(* Logix 5000 project; controller Seperator 1756-L85E rev 33.11; software revision 33.01; part 4 of 7 *)

ADD_ON_INSTRUCTION Random_Izer   (* revision 1.0 *)
VAR_IN_OUT
   Medium_Flash_ON : BOOL; {required}
   Energy : REAL; {required}
END_VAR
VAR_INPUT
   High_Limit_Reached : DINT;
   Actual_To_Same_Interval_Prior_Periods : REAL;
   Production_Lines_To_Like_Lines : REAL;
   Actual_to_Baseline : REAL;
   Production_Runs_To_Like_Runs : REAL;
   Eunits_PER_UOPunits : REAL;
   Edollar_PER_UOPunits : REAL;
   Eunits_PER_UOPdollar : REAL;
   Edollar_PER_UOPdollar : REAL;
   kG_CO2_e : REAL;
   Metric_Tonnes : REAL;
   Water_Demand : REAL;
   Air_Demand : REAL;
   Gas_Demand : REAL;
   Electric_Demand : REAL;
   Steam_Demand : REAL;
   Water_Usage : REAL;
   Air_Usage : REAL;
   Gas_Usage : REAL;
   Electric_Usage : REAL;
   Steam_Usage : REAL;
   work : REAL;
END_VAR
VAR
   APAC_ONS : DINT;
   Low_Limit_Reached : DINT;
   Enable_Low_Check : BOOL; {access None}
   Low_Limit : REAL := 20.0; {access None}
   High_Limit : REAL := 95.0; {access None}
   High_High_Limit : REAL := 100.0; {access None}
   Low_Low_Limit : REAL; {access None}
   Enable_Hi_Check : BOOL; {access None}
   ons1 : BOOL; {access None}
   ons2 : BOOL; {access None}
END_VAR

ROUTINE Logic   (* ladder *)
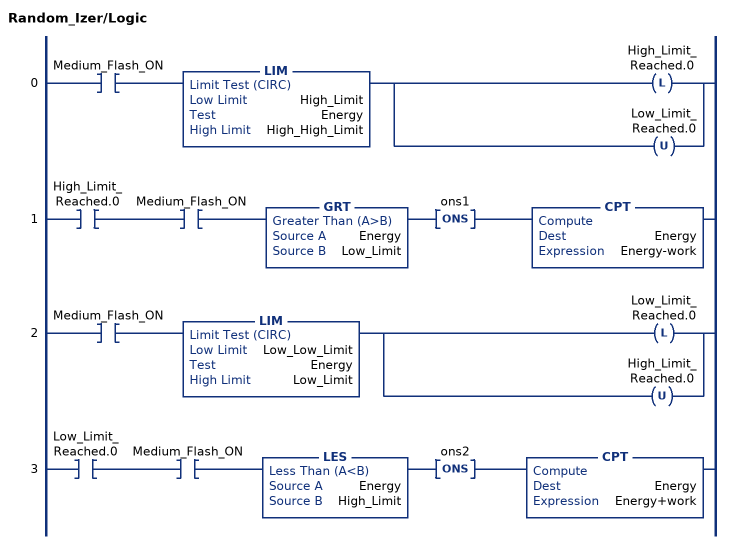
   0: XIC(Medium_Flash_ON)LIM(High_Limit,Energy,High_High_Limit)[OTL(High_Limit_Reached.0) ,OTU(Low_Limit_Reached.0) ];
   1: XIC(High_Limit_Reached.0)XIC(Medium_Flash_ON)GRT(Energy,Low_Limit)ONS(ons1)CPT(Energy,Energy-work);
   2: XIC(Medium_Flash_ON)LIM(Low_Low_Limit,Energy,Low_Limit)[OTL(Low_Limit_Reached.0) ,OTU(High_Limit_Reached.0) ];
   3: XIC(Low_Limit_Reached.0)XIC(Medium_Flash_ON)LES(Energy,High_Limit)ONS(ons2)CPT(Energy,Energy+work);
END_ROUTINE
END_ADD_ON_INSTRUCTION

ADD_ON_INSTRUCTION SineWave   (* revision 1.0, ExecutePrescan *)
VAR_INPUT
   Period : DINT; {visible}
   Max : REAL; {visible}
END_VAR
VAR_IN_OUT
   Out : INT; {required}
END_VAR
VAR
   PI : REAL;
   AlaFillerTimer : TIMER := (PRE := 20000, DN := 1);
   XNum : REAL;
   XDen : REAL;
   Ctrl : CONTROL := (LEN := 1);
   Ctrl2 : CONTROL;
END_VAR

ROUTINE Logic   (* ladder *)
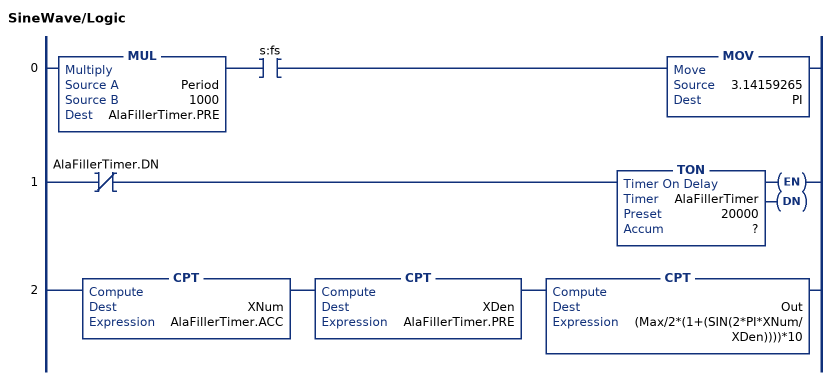
   0: MUL(Period,1000,AlaFillerTimer.PRE)XIC(s:fs)MOV(3.14159265,PI);
   1: XIO(AlaFillerTimer.DN)TON(AlaFillerTimer,?,?);
   2: CPT(XNum,AlaFillerTimer.ACC)CPT(XDen,AlaFillerTimer.PRE)CPT(Out,(Max/2*(1+(SIN(2*PI*XNum/XDen))))*10);
END_ROUTINE

ROUTINE Prescan   (* structured text *)
   Period:=20;
   Max:=50;
END_ROUTINE
END_ADD_ON_INSTRUCTION

ADD_ON_INSTRUCTION UADD   (* revision 1.1, vendor Dr. Frank Jordan / Rockwell Automation *)
// Addition of  two unsigned DINT
// (without overflow / minor faults)
// Revision note:
// This code is provided as application example without any warranty
VAR_INPUT
   V1 : DINT; {visible}
   V2 : DINT; {visible}
END_VAR
VAR_OUTPUT
   Out : DINT; {access Read Only, visible}
   Sts_C : BOOL; {access Read Only, visible}   // Carry result
   Sts_N : BOOL; {access Read Only, visible}   // Negative result
   Sts_V : BOOL; {access Read Only, visible}   // Overflow result
   Sts_Z : BOOL; {access Read Only, visible}   // Zero result
END_VAR
VAR
   V1_Hi : DINT; {access None}
   V1_Lo : DINT; {access None}
   V2_Hi : DINT; {access None}
   V2_Lo : DINT; {access None}
   SumLo : DINT; {access None}
   SumHi : DINT; {access None}
   tmp : DINT; {access None}
END_VAR

ROUTINE Logic   (* ladder *)
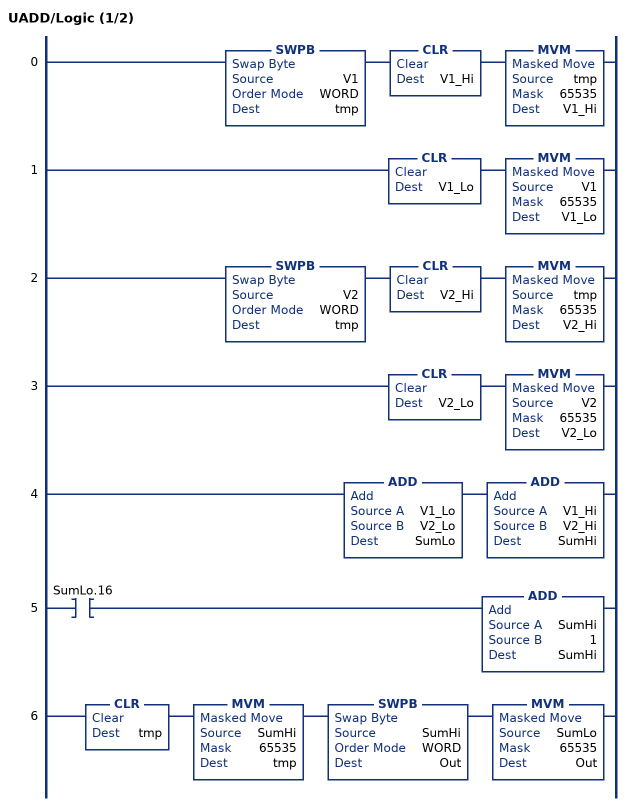
   0: SWPB(V1,WORD,tmp)CLR(V1_Hi)MVM(tmp,65535,V1_Hi);
   1: CLR(V1_Lo)MVM(V1,65535,V1_Lo);
   2: SWPB(V2,WORD,tmp)CLR(V2_Hi)MVM(tmp,65535,V2_Hi);
   3: CLR(V2_Lo)MVM(V2,65535,V2_Lo);
   4: ADD(V1_Lo,V2_Lo,SumLo)ADD(V1_Hi,V2_Hi,SumHi);
   5: XIC(SumLo.16)ADD(SumHi,1,SumHi);
   6: CLR(tmp)MVM(SumHi,65535,tmp)SWPB(SumHi,WORD,Out)MVM(SumLo,65535,Out);
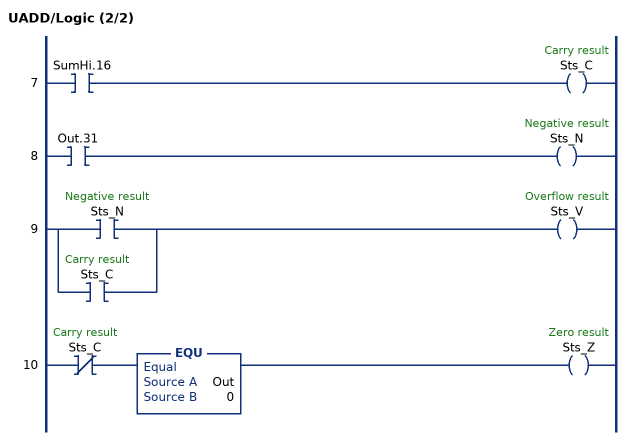
   7: XIC(SumHi.16)OTE(Sts_C);
   8: XIC(Out.31)OTE(Sts_N);
   9: [XIC(Sts_N) ,XIC(Sts_C) ]OTE(Sts_V);
   10: XIO(Sts_C)EQU(Out,0)OTE(Sts_Z);
END_ROUTINE
END_ADD_ON_INSTRUCTION

ADD_ON_INSTRUCTION UMUL   (* revision 1.2, vendor Dr. Frank Jordan / Rockwell Automation *)
// Multiplication of  two unsigned DINT
// (without overflow / minor faults)
// Revision note:
// This code is provided as application example without any warranty
VAR_INPUT
   V1 : DINT; {visible}
   V2 : DINT; {visible}
END_VAR
VAR_OUTPUT
   Sts_C : BOOL; {access Read Only, visible}   // Carry result
   Sts_N : BOOL; {access Read Only, visible}   // Negative result
   Sts_V : BOOL; {access Read Only, visible}   // Overflow result
   Sts_Z : BOOL; {access Read Only, visible}   // Zero result
   Out : DINT; {access Read Only, visible}
END_VAR
VAR
   tmp : DINT; {access None}
   WRK : INT[6]; {access None}
   WRKm : DINT[6]; {access None}
   Low : DINT; {access None}
   Mid : DINT; {access None}
   High : DINT; {access None}
END_VAR

ROUTINE Logic   (* ladder *)
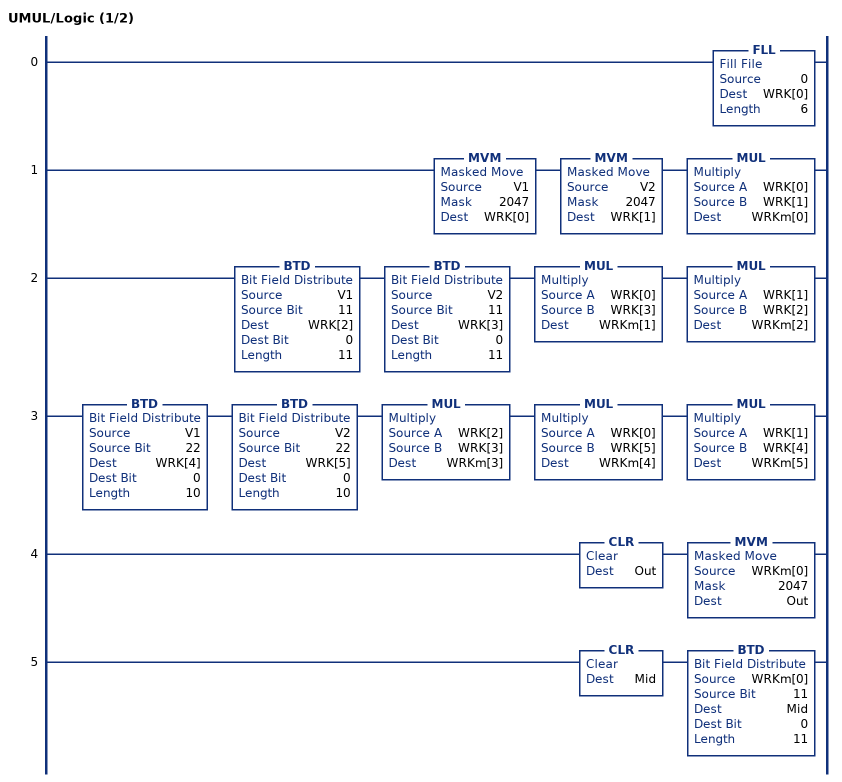
   0: FLL(0,WRK[0],6);
   1: MVM(V1,2047,WRK[0])MVM(V2,2047,WRK[1])MUL(WRK[0],WRK[1],WRKm[0]);
   2: BTD(V1,11,WRK[2],0,11)BTD(V2,11,WRK[3],0,11)MUL(WRK[0],WRK[3],WRKm[1])MUL(WRK[1],WRK[2],WRKm[2]);
   3: BTD(V1,22,WRK[4],0,10)BTD(V2,22,WRK[5],0,10)MUL(WRK[2],WRK[3],WRKm[3])MUL(WRK[0],WRK[5],WRKm[4])MUL(WRK[1],WRK[4],WRKm[5]);
   4: CLR(Out)MVM(WRKm[0],2047,Out);
   5: CLR(Mid)BTD(WRKm[0],11,Mid,0,11);
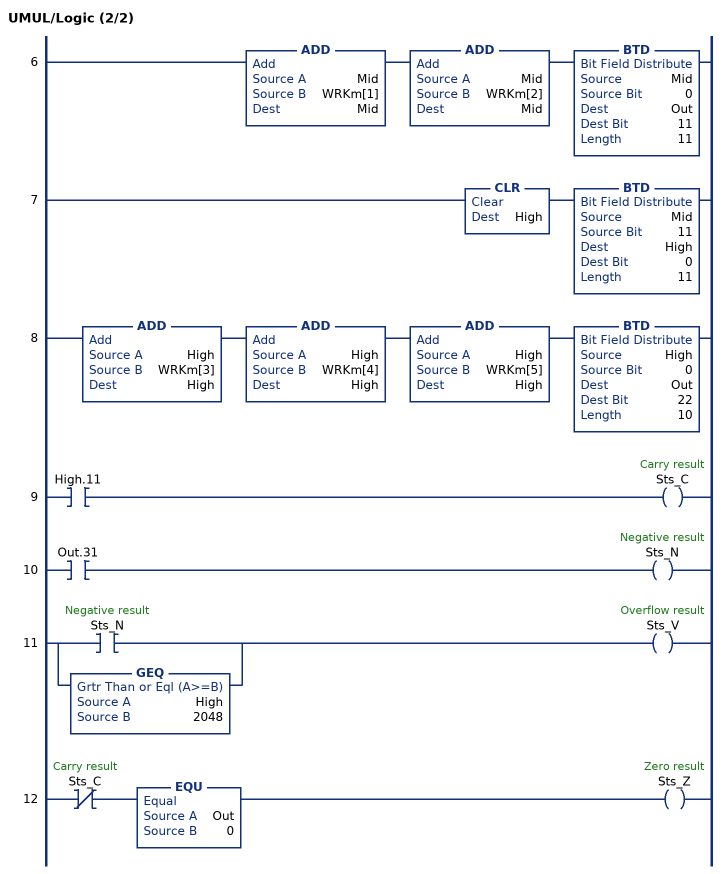
   6: ADD(Mid,WRKm[1],Mid)ADD(Mid,WRKm[2],Mid)BTD(Mid,0,Out,11,11);
   7: CLR(High)BTD(Mid,11,High,0,11);
   8: ADD(High,WRKm[3],High)ADD(High,WRKm[4],High)ADD(High,WRKm[5],High)BTD(High,0,Out,22,10);
   9: XIC(High.11)OTE(Sts_C);
   10: XIC(Out.31)OTE(Sts_N);
   11: [XIC(Sts_N) ,GEQ(High,2048) ]OTE(Sts_V);
   12: XIO(Sts_C)EQU(Out,0)OTE(Sts_Z);
END_ROUTINE
END_ADD_ON_INSTRUCTION

ADD_ON_INSTRUCTION ValveSim   (* revision 1.0, vendor Rockwell, ExecutePrescan *)
VAR_INPUT
   ValveOpenRequest : BOOL;
END_VAR
VAR_OUTPUT
   ValveOpened : BOOL; {access Read Only}
   ValveClosed : BOOL; {access Read Only}
END_VAR
VAR
   OpenCommand : BOOL;
   OpenedCommandDelay : TIMER := (PRE := 1000);
   ClosedCommandDelay : TIMER := (PRE := 1000);
END_VAR

ROUTINE Logic   (* ladder *)
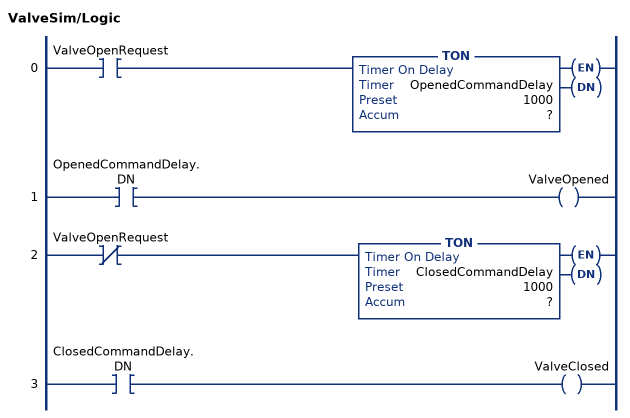
   0: XIC(ValveOpenRequest)TON(OpenedCommandDelay,?,?);
   1: XIC(OpenedCommandDelay.DN)OTE(ValveOpened);
   2: XIO(ValveOpenRequest)TON(ClosedCommandDelay,?,?);
   3: XIC(ClosedCommandDelay.DN)OTE(ValveClosed);
END_ROUTINE

ROUTINE Prescan   (* structured text *)
   OpenedCommandDelay.PRE:=3000;
   ClosedCommandDelay.PRE:=3000;
   
END_ROUTINE
END_ADD_ON_INSTRUCTION

VAR_GLOBAL   (* controller tags *)
   _DriveName_FP : BOOL;
   Aborted : SFC_STEP := (Status := 16#0020_0001, PauseTimer := 1);
   Aborted1 : SFC_STEP := (Status := 16#0020_0001, PauseTimer := 1);
   Aborting : SFC_STEP := (Status := 16#0020_0001, PauseTimer := 1);
   Aborting1 : SFC_STEP := (Status := 16#0020_0001, PauseTimer := 1);
   AE_Digital_Alarm : BOOL := 1;
   Auto_Manual : BOOL := 1;
   batchstrng : STRING := 'Batch ID ';
   bottle_clamp_out_delay : TIMER := (PRE := 1000);
   bottle_clamp_out_delayF1 : TIMER := (PRE := 1000);
   bottle_clamp_out_delayF2 : TIMER := (PRE := 1000);
   bottle_clamp_out_delayF3 : TIMER := (PRE := 1000);
   CAP_clamps_out_Delay : TIMER := (PRE := 1000);
   Capper2_Index_complete : BOOL;
   Capper3_Index_complete : BOOL;
   Capper_Head_Sequencer : DINT := 3;
   Capper_Index_complete : BOOL;
   Capper_Running : BOOL := 1;
   colours : STRING[3] := ([0] := 'Black', [1] := 'Blue', [2] := 'White');
   Comms_OK : BOOL;
   CV1 : REAL := 5000.0;
   CV2 : REAL := 7.0;
   CV3 : DINT := 12;
   Display_number : DINT;
   Equilibrating : SFC_STEP := (Status := 16#0820_0001, DN := 1, PauseTimer := 1, PRE := 5000, T := 5250, TMax := 5250, Count := 1);
   Equilibrating1 : SFC_STEP := (Status := 16#0820_0001, DN := 1, PauseTimer := 1, PRE := 5000, T := 5251, TMax := 5251, Count := 2);
   esd : BOOL;
   Extruder_OEE_Availibility : REAL := 67.5;
   Extruder_OEE_PerfoFillerance : REAL := 59.5;
   Extruder_OEE_Quality : REAL := 89.0;
   Extruder_OEE_Value : REAL := 59.3;
   Extruder_Running : BOOL := 1;
   Extruder_speed_actual : REAL := 161.39124;
   Extruder_speed_SP : DINT := 160;
   FC01 : FTV_ctrl := (nr_of_screens := 5, ActiveScreen := 102, ScreenOverride := 102, delay := 5, Act := 1);
   FI101 : REAL := 10.0;
   FI101_Good_Lower : DINT;
   FI101_Good_Upper : REAL := 2.5;
   FI101_Moving_Analog : Moving_Analog_Indicator := (Value := 10.0, Medium_Alarm := 10.0, High_Alarm := 20.0, Min := 30.0, Max := 40.0);
   FI102 : REAL := 8.0;
   FI102_Good_Lower : REAL := -1.5;
   FI102_Good_Upper : REAL := 1.5;
   FI102_Moving_Analog : Moving_Analog_Indicator := (Value := 8.0, Medium_Alarm := 10.0, High_Alarm := 20.0, Min := 30.0, Max := 40.0);
   Filler2_Index_complete : BOOL;
   Filler3_Index_complete : BOOL;
   Filler_Index_complete : BOOL;
   FillerPUD1 : RampUpDn := (Target := 1000.0, STS_Dn := 1, Time := 5.0, output := 1000.0, CMD_Start := 1);
   FillerPUD2 : RampUpDn := (Target := 5.0, STS_Dn := 1, Time := 5.0, output := 5.0, CMD_Start := 1);
   FillerPUD3 : RampUpDn := (CV := 1000.0, Target := 5000.0, STS_Dn := 1, Time := 5.0, output := 5000.0, CMD_Start := 1);
   FillerPUD4 : RampUpDn := (CV := 5.0, Target := 8.0, STS_Dn := 1, Time := 5.0, output := 8.0, CMD_Start := 1);
   FillerPUD5 : RampUpDn := (CV := 1.0, Target := 10.0, STS_Dn := 1, Time := 5.0, output := 10.0, CMD_Start := 1);
   FillerPUD6 : RampUpDn := (Target := 8.0, STS_Dn := 1, Time := 5.0, output := 8.0, CMD_Start := 1);
   FillerPUD7 : RampUpDn := (CV := 8.0, Target := 12.0, STS_Dn := 1, Time := 5.0, output := 12.0, CMD_Start := 1);
   Filling : SFC_STEP := (Status := 16#0820_0001, DN := 1, PauseTimer := 1, PRE := 5000, T := 5250, TMax := 5250, Count := 1);
   Filling1 : SFC_STEP := (Status := 16#a020_0001, X := 1, SA := 1, PauseTimer := 1, PRE := 5000, T := 3000, TMax := 5249, Count := 3);
   Filling_Nozzle_Down_Delay1 : TIMER := (PRE := 2000);
   Filling_Nozzle_Down_Delay2 : TIMER := (PRE := 2000);
   Filling_Nozzle_Down_Delay3 : TIMER := (PRE := 2000);
   Filling_Nozzle_up_Delay1 : TIMER := (PRE := 1000);
   Filling_Nozzle_up_Delay2 : TIMER := (PRE := 1000);
   Filling_Nozzle_up_Delay3 : TIMER := (PRE := 1000);
   Flushing : SFC_STEP := (Status := 16#0020_0001, PauseTimer := 1, PRE := 10000);
   Flushing1 : SFC_STEP := (Status := 16#0020_0001, PauseTimer := 1, PRE := 10000);
   Half_Sec_PLs : TIMER := (PRE := 500, ACC := 241, EN := 1, TT := 1);
   Head1_Temperature_PID_CV : REAL := 300.0;
   Head1_Temperature_PID_PV : REAL := 175.28792;
   Head1_Temperature_PID_SP : REAL := 180.0;
   Head2_Temperature_PID_CV : REAL := 300.0;
   Head2_Temperature_PID_PV : REAL := 49.0;
   Head2_Temperature_PID_SP : REAL := 176.0;
   Head3_Temperature_PID_CV : REAL := 100.372154;
   Head3_Temperature_PID_PV : REAL := 180.85681;
   Head3_Temperature_PID_SP : REAL := 184.0;
   HMI_Screen_Navigation : DINT;
   HMI_Screen_Navigation1 : INT;
   Holding : SFC_STEP := (Status := 16#0020_0001, PauseTimer := 1);
   Holding1 : SFC_STEP := (Status := 16#0020_0001, PauseTimer := 1);
   Idle : SFC_STEP := (Status := 16#0820_0201, DN := 1, PauseTimer := 1, T := 250, TMax := 250, Count := 1);
   Idle1 : SFC_STEP := (Status := 16#0820_0201, DN := 1, PauseTimer := 1, T := 251, TMax := 251, Count := 3);
   II101 : REAL := 12.0;
   II101_Good_Lower : REAL := -50.0;
   II101_Good_Upper : REAL := 50.0;
   II101_Moving_Analog : Moving_Analog_Indicator := (Value := 12.0, Medium_Alarm := 10.0, High_Alarm := 20.0, Min := 30.0, Max := 40.0);
   Infeed_Pump : P_Motor := (Inp_PermOK := 1, Inp_NBPermOK := 1, Inp_IntlkOK := 1, Inp_NBIntlkOK := 1, Cfg_PCmdClear := 1, Cfg_ProgDefault := 1, Cfg_ShedOnFailToStart := 1, Cfg_ShedOnIOFault := 1, Cfg_HasIntlkTripAlm := 1, Cfg_HasIOFaultAlm := 1, Cfg_FailToStartAckReqd := 1, Cfg_FailToStopAckReqd := 1, Cfg_IntlkTripAckReqd := 1, Cfg_IOFaultAckReqd := 1, Cfg_FailToStartSeverity := 3, Cfg_FailToStopSeverity := 3, Cfg_IntlkTripSeverity := 3, Cfg_IOFaultSeverity := 3, Cfg_SimFdbkT := 2, Cfg_FailToStartT := 10, Cfg_FailToStopT := 10, PCmd_Start := 1, Out_Stop := 1, Val_Cmd := 1, Val_Fdbk := 1, Val_Sts := 7, Val_Mode := 8, Sts_Stopping := 1, Sts_Available := 1, Sts_Prog := 1, Ack_FailToStart := 1, Ack_FailToStop := 1, Ack_IntlkTrip := 1, Ack_IOFault := 1, Rdy_Bypass := 1);
   Led_Code : INT := 3;
   LevelUD1 : RampUpDn := (CV := 95.0, Target := 20.0, STS_RampDown := 1, STS_Ramping := 1, Time := 30.0, output := 52.5, CMD_Start := 1);
   LI101 : REAL := 52.5;
   LI101_Moving_Analog : Moving_Analog_Indicator := (Value := 52.5, Medium_Alarm := 10.0, High_Alarm := 20.0, Min := 30.0, Max := 40.0);
   Logix_Status : Logix_Status_FP := (Set_FaceplateAnimation := 70, Val_ProductCode := 96, MemoryTemp[0] := 5, MemoryTemp[1] := 1, MemoryTemp[3] := -13980, MemoryTemp[4] := 3, MemoryTemp[5] := -4332, MemoryTemp[6] := 125, MemoryTemp[9] := 2, MemoryTemp[11] := -4608, MemoryTemp[12] := 3, MemoryTemp[14] := 128, MemoryTemp[17] := 5, MemoryTemp[21] := 6, MemoryTemp[23] := -14020, MemoryTemp[24] := 3, MemoryTemp[25] := 7, MemoryTemp[27] := -4368, MemoryTemp[28] := 125, Val_raw_data := 12384, Sts_ProductCode := 96, MemoryRequestData[0] := 5, MemoryRequestData[2] := 1, MemoryRequestData[4] := 2, MemoryRequestData[6] := 5, MemoryRequestData[8] := 6, MemoryRequestData[10] := 7, Sts_Run := 1, Sts_Major_fault := 1, Sts_KS_in_remote := 1, Set_Controller_Description := '#10 Mixing Reactor', UpdateDelayTimer.PRE := 1000, UpdateDelayTimer.ACC := 900, UpdateDelayTimer.EN := 1, UpdateDelayTimer.TT := 1, Val_MajorFault.timelow := 158781395, Val_MajorFault.timehigh := 324268, Val_MajorFault.type := 6, Val_MajorFault.code := 1, Val_MajorFault.info[0] := 5, Val_MajorFault.info[1] := 31819, Val_MajorFault.info[2] := 9248, Val_MajorFault.info[3] := -566538954, Val_MFS.timelow := 158781395, Val_MFS.timehigh := 324268, Val_MFS.type := 6, Val_MFS.code := 1, Val_MFS.info[0] := 5, Val_MFS.info[1] := 31819, Val_MFS.info[2] := 9248, Val_MFS.info[3] := -566538954, Sts_IO_LED.Off := 1, Sts_Battery_LED.Off := 1, MemoryData.Free_Mem_IO := 992656, MemoryData.Free_Mem_DT := 33012816, MemoryData.Total_Mem_IO := 1030144, MemoryData.Total_Mem_DT := 33554432, MemoryData.Biggest_IO_Mem_Size_Ava := 992496, MemoryData.Biggest_DT_Mem_Size_Ava := 33012672);
   Main_Sequencer : DINT := 300;
   Main_Sequencer_Emptying : DINT := 220;
   Main_Sequencer_Filling : DINT := 300;
   MC_real : REAL := 200.0;
   Medium_Flash_OFF : TIMER := (PRE := 250, ACC := 129, EN := 1, TT := 1);
   Medium_Flash_ON : TIMER := (PRE := 250, ACC := 251, EN := 1, DN := 1);
   Memory_Message : MESSAGE;
        MessageParameters(ServiceCode := 16#0003, LocalElement := Logix_Status.MemoryRequestData[0], DestinationTag := Logix_Status.MemoryTemp[0], ...)
   ModuleAlaFillerHandshake : BOOL := 1;
   ModuleAlaFillerInProcess : BOOL;
   ModuleAlaFillerName : STRING;
   ModuleAlaFillerTrigger : DINT;
   MyP_Motor : P_Motor := (Inp_RunFdbk := 1, Inp_PermOK := 1, Inp_NBPermOK := 1, Inp_IntlkOK := 1, Inp_NBIntlkOK := 1, Cfg_HasRunFdbk := 1, Cfg_UseRunFdbk := 1, Cfg_HasIntlkObj := 1, Cfg_HasResInhObj := 1, Cfg_HasRunTimeObj := 1, Cfg_PCmdClear := 1, Cfg_ProgDefault := 1, Cfg_ShedOnFailToStart := 1, Cfg_ShedOnIOFault := 1, Cfg_HasFailToStartAlm := 1, Cfg_HasFailToStopAlm := 1, Cfg_HasIntlkTripAlm := 1, Cfg_HasIOFaultAlm := 1, Cfg_FailToStartAckReqd := 1, Cfg_FailToStopAckReqd := 1, Cfg_IntlkTripAckReqd := 1, Cfg_IOFaultAckReqd := 1, Cfg_FailToStartSeverity := 3, Cfg_FailToStopSeverity := 3, Cfg_IntlkTripSeverity := 3, Cfg_IOFaultSeverity := 3, Cfg_SimFdbkT := 15, Cfg_FailToStartT := 10, Cfg_FailToStopT := 10, Out_Run := 1, Val_Fdbk := 1, Val_Sts := 2, Val_Mode := 8, Val_Notify := 1, Sts_Running := 1, Sts_Available := 1, Sts_Prog := 1, Ack_IntlkTrip := 1, Ack_IOFault := 1, Rdy_Bypass := 1, Rdy_ResetAckAll := 1);   // My (Single-Speed, Non-Reversing) Motor
   Operator_Mode : BOOL;
   Phase_Control : Phase_Control;
   Phase_Result : DINT;
   PI102 : REAL := 2.0;
   PI102_Good_Lower : REAL := 0.7;
   PI102_Good_Upper : REAL := 1.3;
   PI102_Moving_Analog : Moving_Analog_Indicator := (Value := 2.0, Medium_Alarm := 10.0, High_Alarm := 20.0, Min := 30.0, Max := 40.0);
   PVP_Init : BOOL;
   Qtr_Sec_PLs : TIMER := (PRE := 250, ACC := 241, EN := 1, TT := 1);
   R1_Head1_Blockage_Sensor : BOOL;
   R1_Head1_Temperature : REAL := 175.28792;
   R1_Head2_Sequencer : DINT := 7;
   R1_Head2_Temperature : REAL := 177.8014;
   R1_Head3_Sequencer : DINT := 7;
   R1_Head3_Temperature : REAL := 180.85681;
   R2_Head1_Blockage_Sensor : BOOL := 1;
   R2_Head1_Sequencer : DINT := 9;
   R2_Head1_Temperature : REAL := 170.32004;
   R2_Head2_Blockage_Sensor : BOOL := 1;
   R2_Head2_Sequencer : DINT := 9;
   R2_Head2_Temperature : REAL := 169.0278;
   R2_Head3_Blockage_Sensor : BOOL := 1;
   R2_Head3_Sequencer : DINT := 9;
   R2_Head3_Temperature : REAL := 170.32004;
   R3_Head1_Blockage_Sensor : BOOL;
   R3_Head1_Sequencer : DINT := 9;
   R3_Head1_Temperature : REAL := 187.06586;
   R3_Head2_Blockage_Sensor : BOOL;
   R3_Head2_Sequencer : DINT := 9;
   R3_Head2_Temperature : REAL := 187.06586;
   R3_Head3_Blockage_Sensor : BOOL;
   R3_Head3_Sequencer : DINT := 9;
   R3_Head3_Temperature : REAL := 187.06586;
   Random : AOI_SIM_RNG_Simple := (Seed := 521288629, Count := 4, Number := 0.03563233);
   Range : DINT := 420;
   Remote_Display_number : DINT;
   Restarting : SFC_STEP := (Status := 16#0020_0001, PauseTimer := 1);
   Restarting1 : SFC_STEP := (Status := 16#0020_0001, PauseTimer := 1);
   Rotary_OEE_Availibility : REAL := 99.94192;
   Rotary_OEE_PerfoFillerance : REAL := 54.122345;
   Rotary_OEE_Quaility : REAL := 98.31933;
   Rotary_OEE_Value : REAL := 86.39993;
   Sec_PLs : TIMER := (PRE := 250, ACC := 237, EN := 1, TT := 1);
   Seperating : SFC_STEP := (Status := 16#0820_0001, DN := 1, PauseTimer := 1, T := 7500, TMax := 7500, Count := 1);
   Seperating1 : SFC_STEP := (Status := 16#0820_0001, DN := 1, PauseTimer := 1, T := 6500, TMax := 7500, Count := 2);
   Seperator_Control : PHASE := (State := 1, Running := 1);
   Seperator_State : BOOL[32] := ([4] := 1);
   Set_Sgl : MESSAGE;
        MessageParameters(ServiceCode := 16#0010, LocalElement := Storage[0], ...)
   Show_AlaFiller_Banner : BOOL;
   Show_AlaFiller_Banner1 : BOOL;
   Show_Capper : BOOL;
   Show_Capper1 : BOOL;
   Show_Capper_Zoom : BOOL;
   Show_Capper_Zoom1 : BOOL;
   Show_Filling_Head : BOOL;
   Show_Filling_Head1 : BOOL;
   Show_Filling_Head_Zoom : BOOL;
   Show_Filling_Head_Zoom1 : BOOL;
   Show_Home : BOOL;
   Show_Home1 : BOOL;
   Show_Network : BOOL;
   Show_Network1 : BOOL;
   Show_Phase_Manager : BOOL;
   Show_Phase_Manager1 : BOOL;
   Show_Separator : BOOL;
   Show_Separator1 : BOOL;
   Show_Tank : BOOL;
   Show_Tank1 : BOOL;
   SP_real : REAL := 61.0;
   Speeding : SFC_STEP := (Status := 16#0820_0001, DN := 1, PauseTimer := 1, T := 9000, TMax := 9000, Count := 1);
   Speeding1 : SFC_STEP := (Status := 16#0820_0001, DN := 1, PauseTimer := 1, T := 6500, TMax := 9000, Count := 2);
   Speeding2 : SFC_STEP := (Status := 16#0820_0001, DN := 1, PauseTimer := 1, T := 6500, TMax := 9000, Count := 2);
   Starting : SFC_STEP := (Status := 16#0820_0001, DN := 1, PauseTimer := 1, T := 7500, TMax := 7500, Count := 1);
   Starting1 : SFC_STEP := (Status := 16#0820_0001, DN := 1, PauseTimer := 1, T := 6500, TMax := 7500, Count := 2);
   Starting2 : SFC_STEP := (Status := 16#0820_0001, DN := 1, PauseTimer := 1, T := 6500, TMax := 7500, Count := 2);
   Startup_Timer_PVP : TIMER := (PRE := 2000);
   Status_Code : INT := 5;
   Status_Code1 : INT := 1;
   Stopped : SFC_STEP := (Status := 16#0020_0001, PauseTimer := 1);
   Stopped1 : SFC_STEP := (Status := 16#0020_0001, PauseTimer := 1);
   Stopped2 : SFC_STEP := (Status := 16#0020_0001, PauseTimer := 1);
   Stopping : SFC_STEP := (Status := 16#0020_0001, PauseTimer := 1);
   Stopping1 : SFC_STEP := (Status := 16#0020_0001, PauseTimer := 1);
   Stopping2 : SFC_STEP := (Status := 16#0020_0001, PauseTimer := 1);
   Storage : SINT[510] := ([0] := 100, [4] := 47, [10] := -68, [11] := -50, [12] := 75, [13] := -28, [14] := -75, [15] := -102, [16] := -76, [17] := 1, [18] := -102, [19] := 13, [20] := 3, [22] := 11, [23] := -21, [24] := 1, [38] := 64, [39] := -37, [40] := -99, [41] := 1, [42] := -103, [43] := -28, [44] := 4, [46] := -19, [47] := 28, [106] := 1, [110] := 2, [111] := 1, [112] := 1, [113] := 1, [114] := 50);
   Storage1 : SINT[510] := ([0] := 100, [4] := 47, [10] := -68, [11] := -50, [12] := 75, [13] := -28, [14] := -75, [15] := -102, [16] := -76, [17] := 1, [18] := -102, [19] := 13, [20] := 3, [22] := 11, [23] := -21, [24] := 1, [38] := 64, [39] := -37, [40] := -99, [41] := 1, [42] := -103, [43] := -28, [44] := 4, [46] := -19, [47] := 28, [106] := 1, [110] := 2, [111] := 1, [112] := 1, [113] := 1, [114] := 50);
   T1 : FBD_TIMER := (TimerEnable := 1, PRE := 15000, ACC := 15000, EN := 1, DN := 1);
   T11 : FBD_TIMER := (TimerEnable := 1, PRE := 15000, ACC := 15000, EN := 1, DN := 1);
   tenfloats : REAL[10] := ([0] := -0.07826284, [1] := 0.09530566, [2] := 0.05149425, [3] := 228.6808, [4] := 0.24815133, [5] := 82.302574);
   TI101 : REAL := 59.672882;
   TI1011 : REAL := 56.0;
   TI101_Good_Lower : REAL := 51.0;
   TI101_Good_Lower1 : REAL := 51.0;
   TI101_Good_Upper : REAL := 61.0;
   TI101_Good_Upper1 : REAL := 61.0;
   TI101_Moving_Analog : Moving_Analog_Indicator := (Value := 59.672882, Medium_Alarm := 10.0, High_Alarm := 20.0, Min := 30.0, Max := 40.0);
   TI101_Temperature : REAL := 281.09085;
   TI101_Temperature_PID_CV : REAL;
   TI101_Temperature_PID_PV : REAL := 59.672882;
   TI101_Temperature_PID_SP : REAL := 56.0;
   VI101 : REAL := 5000.0;
   VI1011 : REAL;
   VI101_Good_Lower : REAL := -50.0;
   VI101_Good_Lower1 : REAL := -50.0;
   VI101_Good_Upper : REAL := 50.0;
   VI101_Good_Upper1 : REAL := 50.0;
   VI101_Moving_Analog : Moving_Analog_Indicator := (Value := 5000.0, Medium_Alarm := 10.0, High_Alarm := 20.0, Min := 30.0, Max := 40.0);
   wct : DINT[2] := ([0] := 3065118, [1] := 322342);
   work : REAL := 0.118;
   work_DINT : DINT := 103;
END_VAR

PROGRAM Capper   (* main routine Initialisation *)
VAR
   autoreset : TIMER := (PRE := 39571);
   autoresetpulse : BOOL;
   batchcountbase : DINT := 35000;
   batchcounter : DINT := 526;
   Capper_Efficiency_FTAE : BOOL[32];
   Capper_Fault_FTAE : BOOL[32];
   Capper_Warning_FTAE : BOOL[32];
   colourcounter : DINT := 1;
   Index_Move : BOOL;
   Index_Move_Timer : TIMER := (PRE := 1000);
   m_slowperc_lim : REAL := 0.92;
   MetricsData : mtrcsdt := (PartId := 'Corner block', IdealCT := 23.7, GoodParts := 13853, ScrapParts := 3717, TotalParts := 17570, Running := 1, Monitored_Availability := 1, Machine_State := 1, BatchID := 'Batch ID 35526', Colour := 'Blue');
   mset_badperc : REAL := 0.07;   // Bad percentage valid: 1.0 - mset_goodperc
   mset_fltfudge : REAL := 0.93;   // fault distribution fudge factor do not change
   mset_fltoffset : DINT := 2;   // fault distribution offset do not change
   mset_goodperc : REAL := 0.85;   // Good percentage valid: 0.51 - 0.99
   mset_wrnfudge : REAL := 0.02;   // warning distribution fudge factor do not change
   mset_wrnoffset : DINT := 2;   // warning distribution offset do not change
   oneshots : DINT;
   tempDINT : DINT := 70;
   tempstring : STRING := '35526';
END_VAR

ROUTINE Capper_Alarms   (* ladder *)
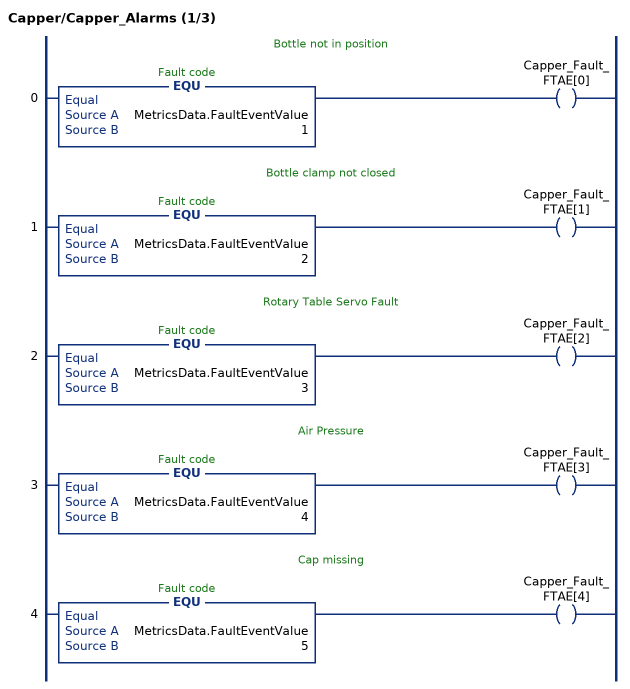
   // Bottle not in position
   0: EQU(MetricsData.FaultEventValue,1)OTE(Capper_Fault_FTAE[0]);
   // Bottle clamp not closed
   1: EQU(MetricsData.FaultEventValue,2)OTE(Capper_Fault_FTAE[1]);
   // Rotary Table Servo Fault
   2: EQU(MetricsData.FaultEventValue,3)OTE(Capper_Fault_FTAE[2]);
   // Air Pressure
   3: EQU(MetricsData.FaultEventValue,4)OTE(Capper_Fault_FTAE[3]);
   // Cap missing
   4: EQU(MetricsData.FaultEventValue,5)OTE(Capper_Fault_FTAE[4]);
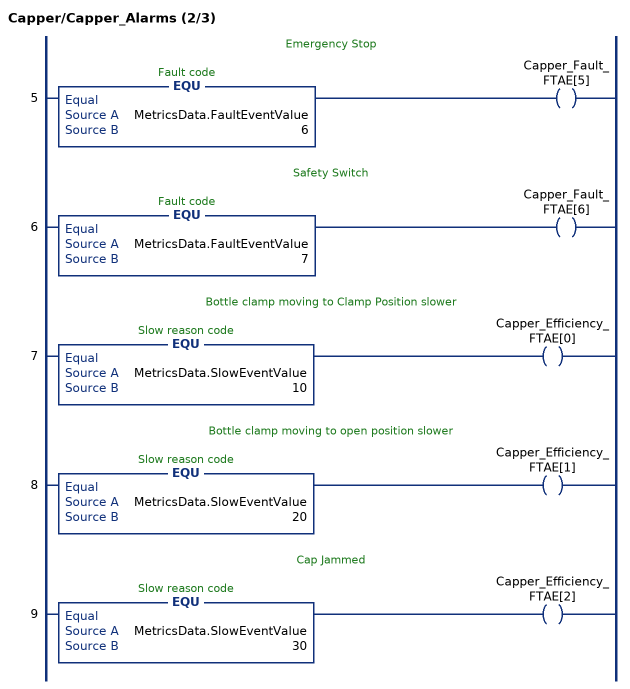
   // Emergency Stop
   5: EQU(MetricsData.FaultEventValue,6)OTE(Capper_Fault_FTAE[5]);
   // Safety Switch
   6: EQU(MetricsData.FaultEventValue,7)OTE(Capper_Fault_FTAE[6]);
   // Bottle clamp moving to Clamp Position slower
   7: EQU(MetricsData.SlowEventValue,10)OTE(Capper_Efficiency_FTAE[0]);
   // Bottle clamp moving to open position slower
   8: EQU(MetricsData.SlowEventValue,20)OTE(Capper_Efficiency_FTAE[1]);
   // Cap Jammed
   9: EQU(MetricsData.SlowEventValue,30)OTE(Capper_Efficiency_FTAE[2]);
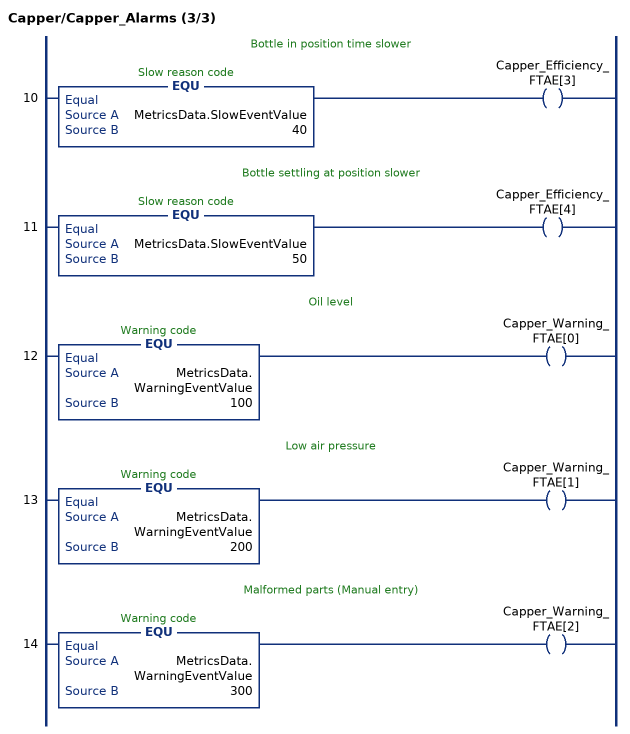
   // Bottle in position time slower
   10: EQU(MetricsData.SlowEventValue,40)OTE(Capper_Efficiency_FTAE[3]);
   // Bottle settling at position slower
   11: EQU(MetricsData.SlowEventValue,50)OTE(Capper_Efficiency_FTAE[4]);
   // Oil level
   12: EQU(MetricsData.WarningEventValue,100)OTE(Capper_Warning_FTAE[0]);
   // Low air pressure
   13: EQU(MetricsData.WarningEventValue,200)OTE(Capper_Warning_FTAE[1]);
   // Malformed parts (Manual entry)
   14: EQU(MetricsData.WarningEventValue,300)OTE(Capper_Warning_FTAE[2]);
END_ROUTINE

ROUTINE Index_Control   (* ladder *)
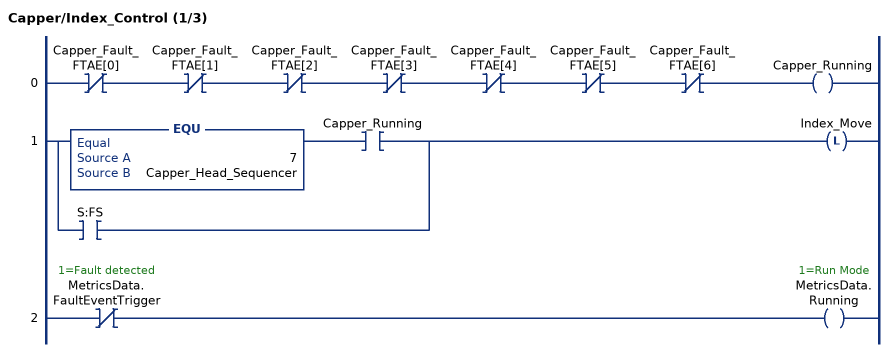
   0: XIO(Capper_Fault_FTAE[0])XIO(Capper_Fault_FTAE[1])XIO(Capper_Fault_FTAE[2])XIO(Capper_Fault_FTAE[3])XIO(Capper_Fault_FTAE[4])XIO(Capper_Fault_FTAE[5])XIO(Capper_Fault_FTAE[6])OTE(Capper_Running);
   1: [EQU(7,Capper_Head_Sequencer) XIC(Capper_Running) ,XIC(S:FS) ]OTL(Index_Move);
   2: XIO(MetricsData.FaultEventTrigger)OTE(MetricsData.Running);
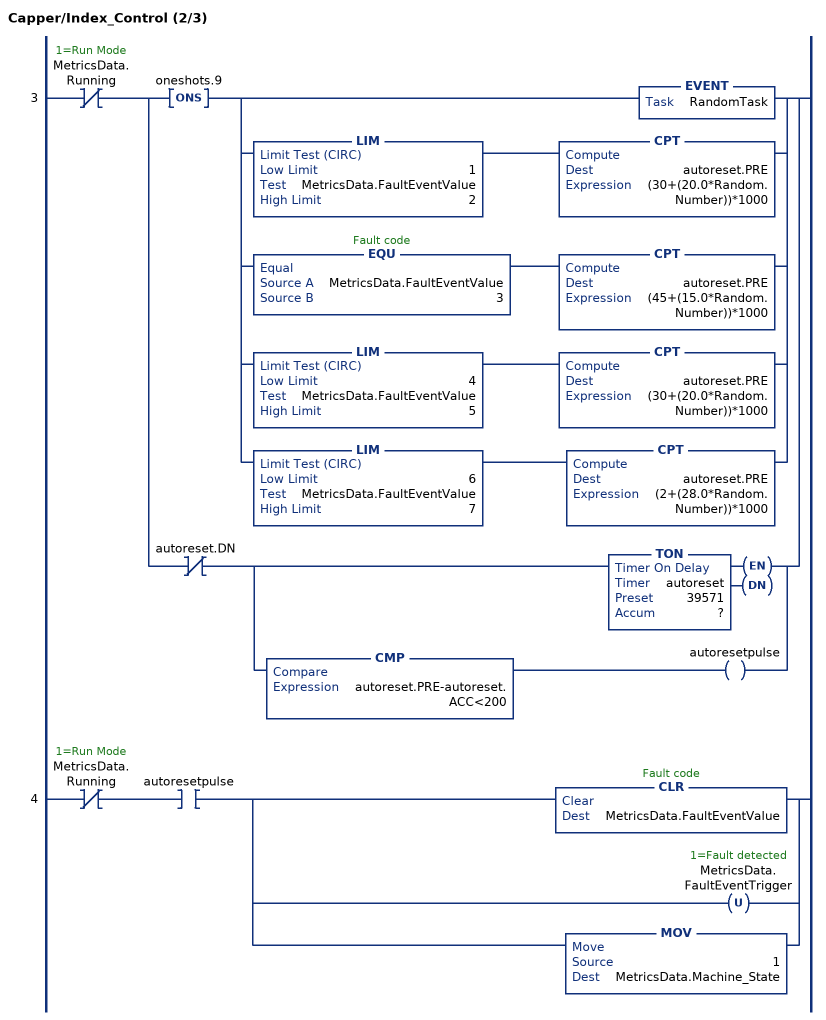
   3: XIO(MetricsData.Running)[ONS(oneshots.9) [EVENT(RandomTask) ,LIM(1,MetricsData.FaultEventValue,2) CPT(autoreset.PRE,(30+(20.0*Random.Number))*1000) ,EQU(MetricsData.FaultEventValue,3) CPT(autoreset.PRE,(45+(15.0*Random.Number))*1000) ,LIM(4,MetricsData.FaultEventValue,5) CPT(autoreset.PRE,(30+(20.0*Random.Number))*1000) ,LIM(6,MetricsData.FaultEventValue,7) CPT(autoreset.PRE,(2+(28.0*Random.Number))*1000) ] ,XIO(autoreset.DN) [TON(autoreset,?,?) ,CMP(autoreset.PRE-autoreset.ACC<200) OTE(autoresetpulse) ] ];
   4: XIO(MetricsData.Running)XIC(autoresetpulse)[CLR(MetricsData.FaultEventValue) ,OTU(MetricsData.FaultEventTrigger) ,MOV(1,MetricsData.Machine_State) ];
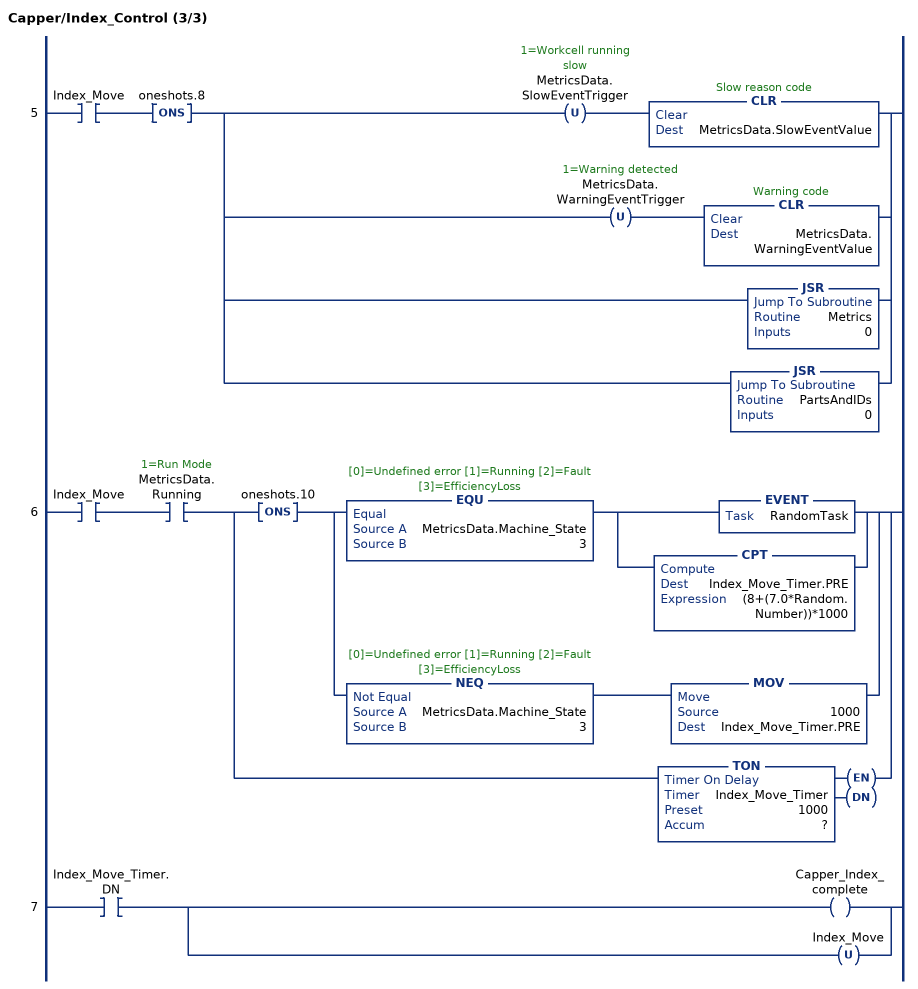
   5: XIC(Index_Move)ONS(oneshots.8)[OTU(MetricsData.SlowEventTrigger) CLR(MetricsData.SlowEventValue) ,OTU(MetricsData.WarningEventTrigger) CLR(MetricsData.WarningEventValue) ,JSR(Metrics,0) ,JSR(PartsAndIDs,0) ];
   6: XIC(Index_Move)XIC(MetricsData.Running)[ONS(oneshots.10) [EQU(MetricsData.Machine_State,3) [EVENT(RandomTask) ,CPT(Index_Move_Timer.PRE,(8+(7.0*Random.Number))*1000) ] ,NEQ(MetricsData.Machine_State,3) MOV(1000,Index_Move_Timer.PRE) ] ,TON(Index_Move_Timer,?,?) ];
   7: XIC(Index_Move_Timer.DN)[OTE(Capper_Index_complete) ,OTU(Index_Move) ];
END_ROUTINE

ROUTINE Initialisation   (* ladder *)
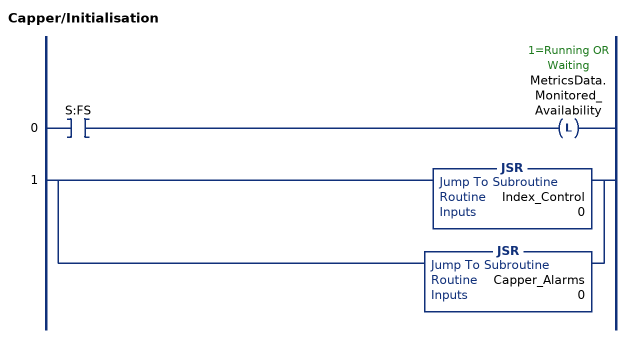
   0: XIC(S:FS)OTL(MetricsData.Monitored_Availability);
   1: [JSR(Index_Control,0) ,JSR(Capper_Alarms,0) ];
END_ROUTINE

ROUTINE Metrics   (* ladder *)
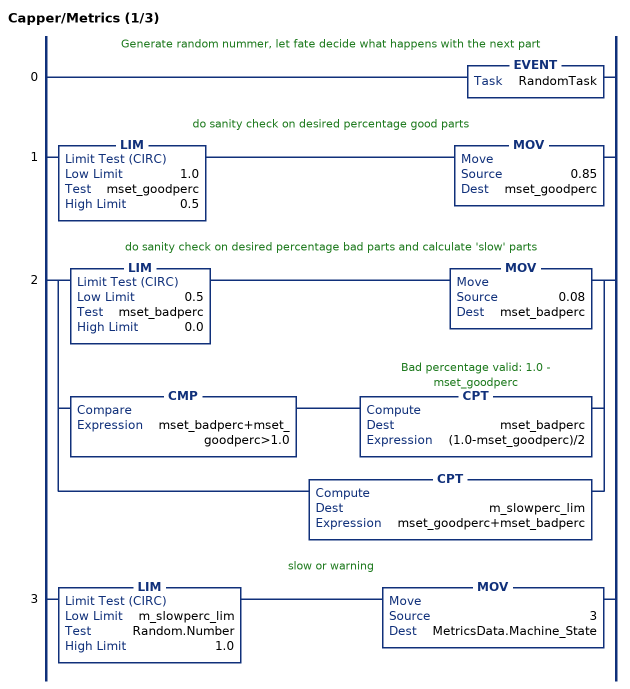
   // Generate random nummer, let fate decide what happens with the next part
   0: EVENT(RandomTask);
   // do sanity check on desired percentage good parts
   1: LIM(1.0,mset_goodperc,0.5)MOV(0.85,mset_goodperc);
   // do sanity check on desired percentage bad parts and calculate 'slow' parts
   2: [LIM(0.5,mset_badperc,0.0) MOV(0.08,mset_badperc) ,CMP(mset_badperc+mset_goodperc>1.0) CPT(mset_badperc,(1.0-mset_goodperc)/2) ,CPT(m_slowperc_lim,mset_goodperc+mset_badperc) ];
   // slow or warning
   3: LIM(m_slowperc_lim,Random.Number,1.0)MOV(3,MetricsData.Machine_State);
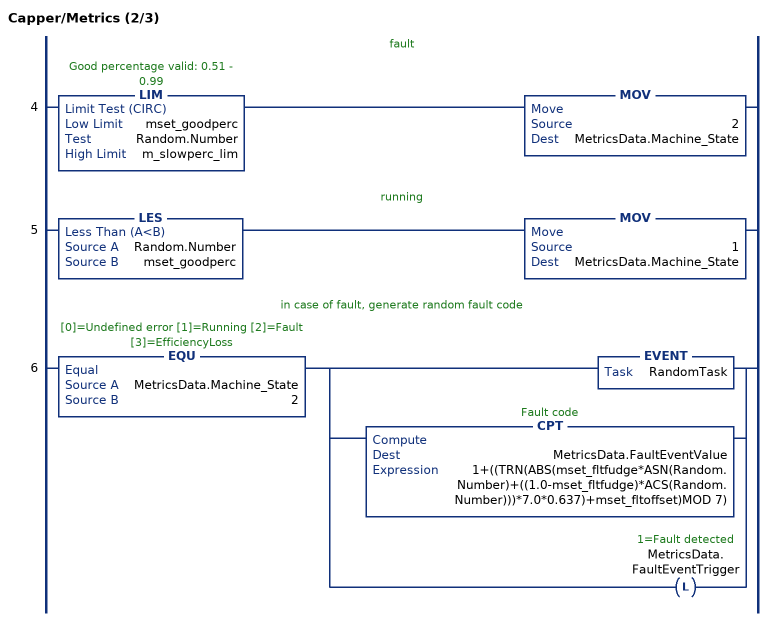
   // fault
   4: LIM(mset_goodperc,Random.Number,m_slowperc_lim)MOV(2,MetricsData.Machine_State);
   // running
   5: LES(Random.Number,mset_goodperc)MOV(1,MetricsData.Machine_State);
   // in case of fault, generate random fault code
   6: EQU(MetricsData.Machine_State,2)[EVENT(RandomTask) ,CPT(MetricsData.FaultEventValue,1+((TRN(ABS(mset_fltfudge*ASN(Random.Number)+((1.0-mset_fltfudge)*ACS(Random.Number)))*7.0*0.637)+mset_fltoffset)MOD 7)) ,OTL(MetricsData.FaultEventTrigger) ];
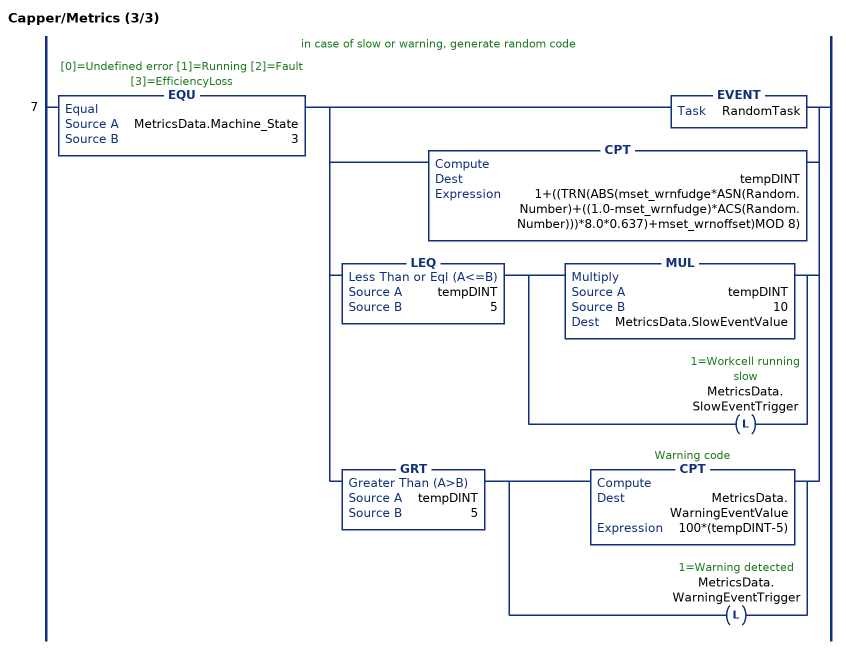
   // in case of slow or warning, generate random code
   7: EQU(MetricsData.Machine_State,3)[EVENT(RandomTask) ,CPT(tempDINT,1+((TRN(ABS(mset_wrnfudge*ASN(Random.Number)+((1.0-mset_wrnfudge)*ACS(Random.Number)))*8.0*0.637)+mset_wrnoffset)MOD 8)) ,LEQ(tempDINT,5) [MUL(tempDINT,10,MetricsData.SlowEventValue) ,OTL(MetricsData.SlowEventTrigger) ] ,GRT(tempDINT,5) [CPT(MetricsData.WarningEventValue,100*(tempDINT-5)) ,OTL(MetricsData.WarningEventTrigger) ] ];
END_ROUTINE

ROUTINE PartsAndIDs   (* ladder *)
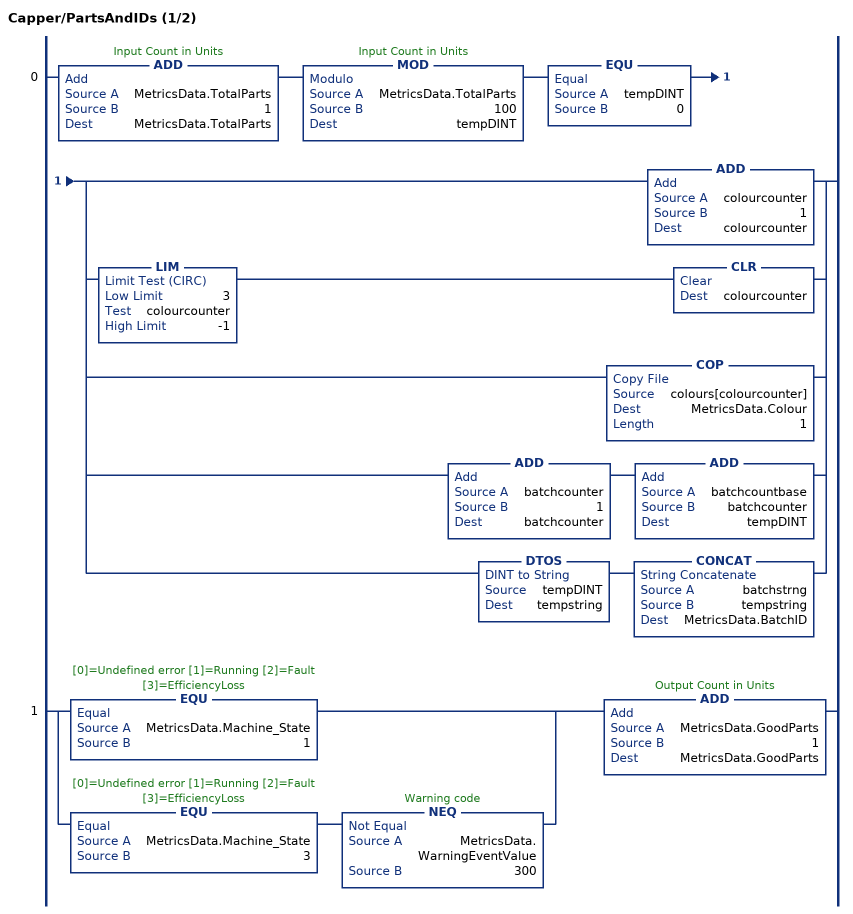
   0: ADD(MetricsData.TotalParts,1,MetricsData.TotalParts)MOD(MetricsData.TotalParts,100,tempDINT)EQU(tempDINT,0)[ADD(colourcounter,1,colourcounter) ,LIM(3,colourcounter,-1) CLR(colourcounter) ,COP(colours[colourcounter],MetricsData.Colour,1) ,ADD(batchcounter,1,batchcounter) ADD(batchcountbase,batchcounter,tempDINT) ,DTOS(tempDINT,tempstring) CONCAT(batchstrng,tempstring,MetricsData.BatchID) ];
   1: [EQU(MetricsData.Machine_State,1) ,EQU(MetricsData.Machine_State,3) NEQ(MetricsData.WarningEventValue,300) ]ADD(MetricsData.GoodParts,1,MetricsData.GoodParts);
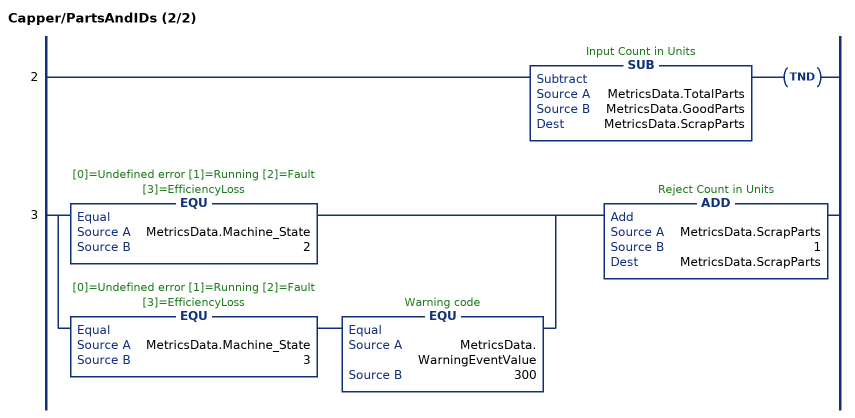
   2: SUB(MetricsData.TotalParts,MetricsData.GoodParts,MetricsData.ScrapParts)TND();
   3: [EQU(MetricsData.Machine_State,2) ,EQU(MetricsData.Machine_State,3) EQU(MetricsData.WarningEventValue,300) ]ADD(MetricsData.ScrapParts,1,MetricsData.ScrapParts);
END_ROUTINE
END_PROGRAM
